FUNCTION "LGF_MatrixSubtraction" : Void   // FC10010, SCL
{ S7_Optimized_Access := 'TRUE' }
   VAR_INPUT
      matrix1 : Array[*, *] of Real;   // minuend
      matrix2 : Array[*, *] of Real;   // subtrahend
   END_VAR
   VAR_OUTPUT
      matrixResult : Array[*, *] of Real;   // result matrix
      error : Bool;
      statusID : UInt;
      status : Word;
   END_VAR
   VAR_TEMP
      tempMatrix1LowerBound1Dim : DInt;   // -
      tempMatrix1LowerBound2Dim : DInt;   // -
      tempMatrix1UpperBound1Dim : DInt;   // -
      tempMatrix1UpperBound2Dim : DInt;   // -
      tempMatrix2LowerBound1Dim : DInt;   // -
      tempMatrix2LowerBound2Dim : DInt;   // -
      tempMatrix2UpperBound1Dim : DInt;   // -
      tempMatrix2UpperBound2Dim : DInt;   // -
      tempResultMatrixLowerBound1Dim : DInt;   // -
      tempResultMatrixLowerBound2Dim : DInt;   // -
      tempResultMatrixUpperBound1Dim : DInt;   // -
      tempResultMatrixUpperBound2Dim : DInt;   // -
      tempCounterDim1 : Int;   // -
      tempCounterDim2 : Int;   // -
   END_VAR
   VAR CONSTANT
      NO_ERROR : Word := 16#0000;   // No errors.
      ERROR_LOWER_BOUND_NOT_EQUAL : Word := 16#8200;   // Lower bounds of matrices are not equal.
      ERROR_UPPER_BOUND_NOT_EQUAL : Word := 16#8201;   // Upper bounds of matrices are not equal.
      ERROR_IN_THIS_BLOCK : UInt := 1;   // statusID: Error in this block.
   END_VAR
BEGIN
   //=============================================================================
   // SIEMENS AG
   // (c)Copyright 2017
   //-----------------------------------------------------------------------------
   // Library:       LGF (Library General Functions)
   // Tested with:   CPU1212C DC/DC/DC FW:V4.2
   // Engineering:   TIA Portal V14 Update 1
   // Restrictions:  -
   // Requirements:  PLC (S7-1200 / S7-1500)
   // Functionality: This function subtracts matrices.
   //-----------------------------------------------------------------------------
   // Change log table:
   // Version  Date        In charge / Changes applied
   // 01.00.00 19.08.2015  Siemens Industry Online Support
   //                      First released version
   // 01.00.01 02.01.2017  Siemens Industry Online Support
   //                      Upgrade: TIA Portal V14 Update 1
   // 02.00.00 06.02.2017  Siemens Industry Online Support
   //                      Functionality using Array[*,*]
   // 02.00.01 17.08.2018  Siemens Industry Online Support
   //                      Upgrade: TIA V15 Update 2
   // 02.00.02 23.11.2018  Siemens Industry Online Support
   //                      Upgrade: TIA V15.1
   //=============================================================================

   //Set "No error" status
   #error := false;
   #statusID := #ERROR_IN_THIS_BLOCK;
   #status := #NO_ERROR;

   // Init resultMatrix
   #matrixResult[0, 0] := 0.0;

   //Determine the size of the matrices
   // Lower bound dimension 1
   #tempMatrix1LowerBound1Dim := LOWER_BOUND(ARR := #matrix1, DIM := 1);
   #tempMatrix2LowerBound1Dim := LOWER_BOUND(ARR := #matrix2, DIM := 1);
   #tempResultMatrixLowerBound1Dim := LOWER_BOUND(ARR := #matrixResult, DIM := 1);
   // Lower bound dimension 2
   #tempMatrix1LowerBound2Dim := LOWER_BOUND(ARR := #matrix1, DIM := 2);
   #tempMatrix2LowerBound2Dim := LOWER_BOUND(ARR := #matrix2, DIM := 2);
   #tempResultMatrixLowerBound2Dim := LOWER_BOUND(ARR := #matrixResult, DIM := 2);
   // Upper bound dimension 1
   #tempMatrix1UpperBound1Dim := UPPER_BOUND(ARR := #matrix1, DIM := 1);
   #tempMatrix2UpperBound1Dim := UPPER_BOUND(ARR := #matrix2, DIM := 1);
   #tempResultMatrixUpperBound1Dim := UPPER_BOUND(ARR := #matrixResult, DIM := 1);
   // Upper bound dimension 2
   #tempMatrix1UpperBound2Dim := UPPER_BOUND(ARR := #matrix1, DIM := 2);
   #tempMatrix2UpperBound2Dim := UPPER_BOUND(ARR := #matrix2, DIM := 2);
   #tempResultMatrixUpperBound2Dim := UPPER_BOUND(ARR := #matrixResult, DIM := 2);

   // Check the lower bound of all matrices
   IF (#tempMatrix1LowerBound1Dim <> #tempMatrix2LowerBound1Dim) OR (#tempMatrix1LowerBound1Dim <> #tempResultMatrixLowerBound1Dim) OR
     (#tempMatrix1LowerBound2Dim <> #tempMatrix2LowerBound2Dim) OR (#tempMatrix1LowerBound2Dim <> #tempResultMatrixLowerBound2Dim) THEN
     #error := TRUE;
     #status := #ERROR_LOWER_BOUND_NOT_EQUAL;
     RETURN;
   END_IF;
   // Check the upper bound of all matrices
   IF (#tempMatrix1UpperBound1Dim <> #tempMatrix2UpperBound1Dim) OR (#tempMatrix1UpperBound1Dim <> #tempResultMatrixUpperBound1Dim) OR
     (#tempMatrix1UpperBound2Dim <> #tempMatrix2UpperBound2Dim) OR (#tempMatrix1UpperBound2Dim <> #tempResultMatrixUpperBound2Dim) THEN
     #error := TRUE;
     #status := #ERROR_UPPER_BOUND_NOT_EQUAL;
     RETURN;
   END_IF;

   // Subtraction of two matrices
   FOR #tempCounterDim1 := #tempMatrix1LowerBound1Dim TO #tempMatrix1UpperBound1Dim DO
     FOR #tempCounterDim2 := #tempMatrix1LowerBound2Dim TO #tempMatrix1UpperBound2Dim DO
       #matrixResult[#tempCounterDim1, #tempCounterDim2] := #matrix1[#tempCounterDim1, #tempCounterDim2] - #matrix2[#tempCounterDim1, #tempCounterDim2];
     END_FOR;
   END_FOR;
END_FUNCTION

FUNCTION "LGF_MatrixTranspose" : Void   // FC10011, SCL
{ S7_Optimized_Access := 'TRUE' }
   VAR_INPUT
      matrix : Array[*, *] of Real;   // Matrix to be transposed.
   END_VAR
   VAR_OUTPUT
      matrixResult : Array[*, *] of Real;   // Transposed matrix.
      error : Bool;
      statusID : UInt;
      status : Word;
   END_VAR
   VAR_TEMP
      tempMatrixLowerBound1Dim : DInt;   // -
      tempMatrixLowerBound2Dim : DInt;   // -
      tempMatrixUpperBound1Dim : DInt;   // -
      tempMatrixUpperBound2Dim : DInt;   // -
      tempResultMatrixLowerBound1Dim : DInt;   // -
      tempResultMatrixLowerBound2Dim : DInt;   // -
      tempResultMatrixUpperBound1Dim : DInt;   // -
      tempResultMatrixUpperBound2Dim : DInt;   // -
      tempCounterDim1 : Int;   // -
      tempCounterDim2 : Int;   // -
   END_VAR
   VAR CONSTANT
      NO_ERROR : Word := 16#0000;   // No error.
      ERROR_LOWER_BOUND : Word := 16#8200;   // Lower bound of "matrixResult" is different to "matrix".
      ERROR_UPPER_BOUND : Word := 16#8201;   // Upper bound of "matrixResult" is different to "matrix".
      ERROR_IN_THIS_BLOCK : UInt := 1;   // statusID: Error in this block.
   END_VAR
BEGIN
   //=============================================================================
   // SIEMENS AG
   // (c)Copyright 2017
   //-----------------------------------------------------------------------------
   // Library:       LGF (Library General Functions)
   // Tested with:   CPU1212C DC/DC/DC FW:V4.2
   // Engineering:   TIA Portal V14 Update 1
   // Restrictions:  -
   // Requirements:  PLC (S7-1200 / S7-1500)
   // Functionality: This function transposes matrices.
   //-----------------------------------------------------------------------------
   // Change log table:
   // Version  Date        In charge / Changes applied
   // 01.00.00 19.08.2015  Siemens Industry Online Support
   //                      First released version
   // 01.00.01 02.01.2017  Siemens Industry Online Support
   //                      Upgrade: TIA Portal V14 Update 1
   // 02.00.00 06.02.2017  Siemens Industry Online Support
   //                      Functionality using Array[*,*]
   // 02.00.01 17.08.2018  Siemens Industry Online Support
   //                      Upgrade: TIA V15 Update 2
   // 02.00.02 23.11.2018  Siemens Industry Online Support
   //                      Upgrade: TIA V15.1
   //=============================================================================

   //Set "No error" status
   #error := false;
   #statusID := #ERROR_IN_THIS_BLOCK;
   #status := #NO_ERROR;

   // Init resultMatrix
   #matrixResult[0, 0] := 0.0;

   //Determine the size of the matrices
   // Lower bound dimension 1
   #tempMatrixLowerBound1Dim := LOWER_BOUND(ARR := #matrix, DIM := 1);
   #tempResultMatrixLowerBound1Dim := LOWER_BOUND(ARR := #matrixResult, DIM := 1);
   // Lower bound dimension 2
   #tempMatrixLowerBound2Dim := LOWER_BOUND(ARR := #matrix, DIM := 2);
   #tempResultMatrixLowerBound2Dim := LOWER_BOUND(ARR := #matrixResult, DIM := 2);
   // Upper bound dimension 1
   #tempMatrixUpperBound1Dim := UPPER_BOUND(ARR := #matrix, DIM := 1);
   #tempResultMatrixUpperBound1Dim := UPPER_BOUND(ARR := #matrixResult, DIM := 1);
   // Upper bound dimension 2
   #tempMatrixUpperBound2Dim := UPPER_BOUND(ARR := #matrix, DIM := 2);
   #tempResultMatrixUpperBound2Dim := UPPER_BOUND(ARR := #matrixResult, DIM := 2);

   // Check whether lower bounds of "matrixResult suit to the input "matrix"
   IF (#tempMatrixLowerBound1Dim <> #tempResultMatrixLowerBound2Dim) OR (#tempMatrixLowerBound2Dim <> #tempResultMatrixLowerBound1Dim) THEN
     #error := TRUE;
     #status := #ERROR_LOWER_BOUND;
     RETURN;
   END_IF;
   // Check whether upper bounds of "matrixResult suit to the input "matrix"
   IF (#tempMatrixUpperBound1Dim <> #tempResultMatrixUpperBound2Dim) OR (#tempMatrixUpperBound2Dim <> #tempResultMatrixUpperBound1Dim) THEN
     #error := TRUE;
     #status := #ERROR_UPPER_BOUND;
     RETURN;
   END_IF;

   //Transpose of the matrix
   FOR #tempCounterDim1 := #tempMatrixLowerBound1Dim TO #tempMatrixUpperBound1Dim DO
     FOR #tempCounterDim2 := #tempMatrixLowerBound2Dim TO #tempMatrixUpperBound2Dim DO
       #matrixResult[#tempCounterDim2, #tempCounterDim1] := #matrix[#tempCounterDim1, #tempCounterDim2];
     END_FOR;
   END_FOR;
END_FUNCTION

FUNCTION "LGF_RandomReal" : Real   // FC10014, SCL
{ S7_Optimized_Access := 'TRUE' }
   VAR_INPUT
      minValue : Real;   // minimal Value random can reach
      maxValue : Real;   // maximal Value random can reach
   END_VAR
   VAR_OUTPUT
      error : Bool;
      statusID : UInt;
      status : Word;
   END_VAR
   VAR_TEMP
      tempTime : DTL;
      tempTimeStatus : Int;
      tempRandomValue : UDInt;
      tempNormReal : Real;
   END_VAR
   VAR CONSTANT
      NO_ERROR : Word := 16#0000;
      NO_CURRENT_JOBS : Word := 16#7000;
      MAX_LESS_MIN : Word := 16#8200;
      ERROR_IN_THIS_BLOCK : UInt := 1;
      ERROR_RD_SYS_T : UInt := 2;
      MIN_UDINT : UDInt := 0;
      MAX_UDINT : UDInt := 4294967295;
   END_VAR
BEGIN
   //=============================================================================
   // Siemens AG
   // (c)Copyright 2017
   //-----------------------------------------------------------------------------
   // Library:       LGF (Library General Functions)
   // Tested with:   CPU1212C DC/DC/DC FW:V4.2
   // Engineering:   TIA Portal V14 Update 1
   // Restrictions:  -
   // Requirements:  PLC (S7-1200 / S7-1500)
   // Functionality: This function generates random numbers in defined limits
   //                (Datatype Real)
   //-----------------------------------------------------------------------------
   // Change log table:
   // Version  Date        In charge / Changes applied
   // 01.00.00 19.08.2015  Siemens Industry Online Support
   //                      First released version
   // 01.00.01 02.01.2017  Siemens Industry Online Support
   //                      Upgrade: TIA Portal V14 Update 1
   // 01.00.02 02.03.2017  Siemens Industry Online Support
   //                      Bugfix: FC number
   // 01.00.03 17.08.2018  Siemens Industry Online Support
   //                      Upgrade: TIA V15 Update 2
   // 01.00.04 23.11.2018  Siemens Industry Online Support
   //                      Upgrade: TIA V15.1
   //-----------------------------------------------------------------------------
   //Status Codes:
   // 16#7000:  No current jobs
   // 16#0000:  Job finished   // Note: There is no "Busy"-Status because the
   //           block is finished within a single cycle
   // 16#8200:  maxValue is samller then minValue 
   //=============================================================================

   //Set "No current job" status
   #error := false;
   #statusID := #ERROR_IN_THIS_BLOCK;
   #status := #NO_CURRENT_JOBS;

   //Check if the maximal Value is less than the minimal value
   IF (#minValue > #maxValue) THEN
     #error := true;
     #statusID := #ERROR_IN_THIS_BLOCK;
     #status := #MAX_LESS_MIN;
     #LGF_RandomReal := 0;
     RETURN;
   END_IF;

   //Read system time
   #tempTimeStatus := RD_SYS_T(#tempTime);

   IF (#tempTimeStatus <> 0) THEN
     #error := true;
     #statusID := #ERROR_RD_SYS_T;
     #status := INT_TO_WORD(#tempTimeStatus);
     #LGF_RandomReal := 0;
     RETURN;
   END_IF;

   //Callculate a random-start-value depending on the time
   #tempRandomValue.%B3 := #tempTime.NANOSECOND.%B0;
   #tempRandomValue.%B2 := #tempTime.NANOSECOND.%B1;
   #tempRandomValue.%B1 := #tempTime.NANOSECOND.%B2;
   #tempRandomValue.%B0 := #tempTime.NANOSECOND.%B3;

   //adapt the calculated random number to the given number span
   #tempNormReal := NORM_X(MIN := #MIN_UDINT, VALUE := #tempRandomValue, MAX := #MAX_UDINT);
   #LGF_RandomReal := SCALE_X(MIN := #minValue, VALUE := #tempNormReal, MAX := #maxValue);

   #status := #NO_ERROR;
END_FUNCTION

FUNCTION "LGF_SearchMinMax" : Void   // FC10015, SCL
{ S7_Optimized_Access := 'TRUE' }
   VAR_INPUT
      variableArray : Variant;
   END_VAR
   VAR_OUTPUT
      minValue : Variant;
      minArrayIndex : Int;
      maxValue : Variant;
      maxArrayIndex : Int;
      error : Bool;
      statusID : UInt;
      status : Word;
   END_VAR
   VAR_TEMP
      tempArraySize : UDInt;
      tempSizeCounter : Int;
      tempInternalError : Int;
      tempActValueInt : Int;
      tempMinInt : Int;
      tempArrayIndexMin : Int;
      tempMaxInt : Int;
      tempArrayIndexMax : Int;
      tempActValueUInt : UInt;
      tempMinUInt : UInt;
      tempMaxUInt : UInt;
      tempActValueDInt : DInt;
      tempMinDInt : DInt;
      tempMaxDInt : DInt;
      tempActValueUDInt : UDInt;
      tempMinUDInt : UDInt;
      tempMaxUDInt : UDInt;
      tempActValueUSInt : USInt;
      tempMinUSInt : USInt;
      tempMaxUSInt : USInt;
      tempActValueSInt : SInt;
      tempMinSInt : SInt;
      tempMaxSInt : SInt;
      tempActValueReal : Real;
      tempMinReal : Real;
      tempMaxReal : Real;
   END_VAR
   VAR CONSTANT
      NO_ERROR : Word := 16#0000;
      NO_CURRENT_JOBS : Word := 16#7000;
      NO_ARRAY : Word := 16#8200;
      WRONG_TYPE : Word := 16#8201;
      NOT_EQUAL_TYPES : Word := 16#8202;
      ERROR_IN_THIS_BLOCK : UInt := 1;
      ERROR_MOVE_BLK_VARIANT : UInt := 2;
   END_VAR
BEGIN
   //=============================================================================
   // SIEMENS AG
   // (c)Copyright 2017
   //-----------------------------------------------------------------------------
   // Library:       LGF (Library General Functions)
   // Tested with:   CPU1212C DC/DC/DC FW:V4.2
   // Engineering:   TIA Portal V14 Update 1
   // Restrictions:  -
   // Requirements:  PLC (S7-1200 / S7-1500)
   // Functionality: This function searches the min and max value in an array
   //-----------------------------------------------------------------------------
   // Change log table:
   // Version  Date        In charge / Changes applied
   // 01.00.00 19.08.2015  Siemens Industry Online Support
   //                      First released version
   // 01.00.01 02.01.2017  Siemens Industry Online Support
   //                      Upgrade: TIA Portal V14 Update 1
   // 01.00.02 17.08.2018  Siemens Industry Online Support
   //                      Upgrade: TIA V15 Update 2
   // 01.00.03 23.11.2018  Siemens Industry Online Support
   //                      Upgrade: TIA V15.1
   //=============================================================================

   // Set "No current job" status
   #error := false;
   #statusID := #ERROR_IN_THIS_BLOCK;
   #status := #NO_CURRENT_JOBS;
   #tempInternalError := 0;

   // Check if the variant-variable is an array if yes cout the elements of the array
   IF NOT (IS_ARRAY(#variableArray)) THEN
     #error := true;
     #statusID := #ERROR_IN_THIS_BLOCK;
     #status := #NO_ARRAY;
     RETURN;
   ELSE
     #tempArraySize := CountOfElements(#variableArray);
   END_IF;

   // Check if the elements of the array and the variables min and max have the same datatype.
   IF TypeOfElements(#variableArray) <> TypeOf(#minValue) OR TypeOf(#minValue) <> TypeOf(#maxValue) THEN
     #error := true;
     #statusID := #ERROR_IN_THIS_BLOCK;
     #status := #NOT_EQUAL_TYPES;
     RETURN;
   END_IF;

   //Request of the datatype
   CASE TypeOfElements(#variableArray) OF
     Int:
       //----------------------- Search min -------------------------------
       #tempMinInt := 32767;
       FOR #tempSizeCounter := 0 TO UDINT_TO_INT(#tempArraySize) DO

         //Read the next element of the array
         #tempInternalError := MOVE_BLK_VARIANT(SRC := #variableArray,
                                                COUNT := 1,
                                                SRC_INDEX := #tempSizeCounter,
                                                DEST_INDEX := 0,
                                                DEST => #tempActValueInt);

         //compare the new value with the actual best value
         IF #tempActValueInt < #tempMinInt THEN
           #tempMinInt := #tempActValueInt;
           #tempArrayIndexMin := #tempSizeCounter;
         END_IF;

       END_FOR;

       //copy the data to the outputs
       #minArrayIndex := #tempArrayIndexMin;
       #tempInternalError := MOVE_BLK_VARIANT(SRC := #tempMinInt,
                                              COUNT := 1,
                                              SRC_INDEX := 0,
                                              DEST_INDEX := 0,
                                              DEST => #minValue);

       //----------------------- Search max -------------------------------
       #tempMaxInt := -32768;
       FOR #tempSizeCounter := 0 TO UDINT_TO_INT(#tempArraySize) DO

         //Read the next element of the array
         #tempInternalError := MOVE_BLK_VARIANT(SRC := #variableArray,
                                                COUNT := 1,
                                                SRC_INDEX := #tempSizeCounter,
                                                DEST_INDEX := 0,
                                                DEST => #tempActValueInt);

         //compare the new value with the actual best value
         IF #tempActValueInt > #tempMaxInt THEN
           #tempMaxInt := #tempActValueInt;
           #tempArrayIndexMax := #tempSizeCounter;
         END_IF;

       END_FOR;

       //copy the data to the outputs
       #maxArrayIndex := #tempArrayIndexMax;
       #tempInternalError := MOVE_BLK_VARIANT(SRC := #tempMaxInt,
                                              COUNT := 1,
                                              SRC_INDEX := 0,
                                              DEST_INDEX := 0,
                                              DEST => #maxValue);

     UInt:
       //----------------------- Search min -------------------------------
       #tempMinUInt := 65535;
       FOR #tempSizeCounter := 0 TO UDINT_TO_INT(#tempArraySize) DO

         //Read the next element of the array
         #tempInternalError := MOVE_BLK_VARIANT(SRC := #variableArray,
                                                COUNT := 1,
                                                SRC_INDEX := #tempSizeCounter,
                                                DEST_INDEX := 0,
                                                DEST => #tempActValueUInt);

         //compare the new value with the actual best value
         IF #tempActValueUInt < #tempMinUInt THEN
           #tempMinUInt := #tempActValueUInt;
           #tempArrayIndexMin := #tempSizeCounter;
         END_IF;

       END_FOR;

       //copy the data to the outputs
       #minArrayIndex := #tempArrayIndexMin;
       #tempInternalError := MOVE_BLK_VARIANT(SRC := #tempMinUInt,
                                              COUNT := 1,
                                              SRC_INDEX := 0,
                                              DEST_INDEX := 0,
                                              DEST => #minValue);

       //----------------------- Search max -------------------------------
       #tempMaxUInt := 0;
       FOR #tempSizeCounter := 0 TO UDINT_TO_INT(#tempArraySize) DO

         //Read the next element of the array
         #tempInternalError := MOVE_BLK_VARIANT(SRC := #variableArray,
                                                COUNT := 1,
                                                SRC_INDEX := #tempSizeCounter,
                                                DEST_INDEX := 0,
                                                DEST => #tempActValueUInt);

         //compare the new value with the actual best value
         IF #tempActValueUInt > #tempMaxUInt THEN
           #tempMaxUInt := #tempActValueUInt;
           #tempArrayIndexMax := #tempSizeCounter;
         END_IF;

       END_FOR;

       //copy the data to the outputs
       #maxArrayIndex := #tempArrayIndexMax;
       #tempInternalError := MOVE_BLK_VARIANT(SRC := #tempMaxUInt,
                                              COUNT := 1,
                                              SRC_INDEX := 0,
                                              DEST_INDEX := 0,
                                              DEST => #maxValue);

     DInt:
       //----------------------- Search min -------------------------------
       #tempMinDInt := 2147483647;
       FOR #tempSizeCounter := 0 TO UDINT_TO_INT(#tempArraySize) DO

         #tempInternalError := MOVE_BLK_VARIANT(SRC := #variableArray,
                                                COUNT := 1,
                                                SRC_INDEX := #tempSizeCounter,
                                                DEST_INDEX := 0,
                                                DEST => #tempActValueDInt);
         IF #tempActValueDInt < #tempMinDInt THEN
           #tempMinDInt := #tempActValueDInt;
           #tempArrayIndexMin := #tempSizeCounter;
         END_IF;

       END_FOR;

       #minArrayIndex := #tempArrayIndexMin;
       #tempInternalError := MOVE_BLK_VARIANT(SRC := #tempMinDInt,
                                              COUNT := 1,
                                              SRC_INDEX := 0,
                                              DEST_INDEX := 0,
                                              DEST => #minValue);

       //----------------------- Search max -------------------------------
       #tempMaxDInt := -2147483648;
       FOR #tempSizeCounter := 0 TO UDINT_TO_INT(#tempArraySize) DO

         #tempInternalError := MOVE_BLK_VARIANT(SRC := #variableArray,
                                                COUNT := 1,
                                                SRC_INDEX := #tempSizeCounter,
                                                DEST_INDEX := 0,
                                                DEST => #tempActValueDInt);
         IF #tempActValueDInt > #tempMaxDInt THEN
           #tempMaxDInt := #tempActValueDInt;
           #tempArrayIndexMax := #tempSizeCounter;
         END_IF;

       END_FOR;

       #maxArrayIndex := #tempArrayIndexMax;
       #tempInternalError := MOVE_BLK_VARIANT(SRC := #tempMaxDInt,
                                              COUNT := 1,
                                              SRC_INDEX := 0,
                                              DEST_INDEX := 0,
                                              DEST => #maxValue);

     UDInt:
       //----------------------- Search min -------------------------------
       #tempMinUDInt := 4294967295;
       FOR #tempSizeCounter := 0 TO UDINT_TO_INT(#tempArraySize) DO

         #tempInternalError := MOVE_BLK_VARIANT(SRC := #variableArray,
                                                COUNT := 1,
                                                SRC_INDEX := #tempSizeCounter,
                                                DEST_INDEX := 0,
                                                DEST => #tempActValueUDInt);
         IF #tempActValueUDInt < #tempMinUDInt THEN
           #tempMinUDInt := #tempActValueUDInt;
           #tempArrayIndexMin := #tempSizeCounter;
         END_IF;

       END_FOR;

       #minArrayIndex := #tempArrayIndexMin;
       #tempInternalError := MOVE_BLK_VARIANT(SRC := #tempMinUDInt,
                                              COUNT := 1,
                                              SRC_INDEX := 0,
                                              DEST_INDEX := 0,
                                              DEST => #minValue);

       //----------------------- Search max -------------------------------
       #tempMaxUDInt := 0;
       FOR #tempSizeCounter := 0 TO UDINT_TO_INT(#tempArraySize) DO

         #tempInternalError := MOVE_BLK_VARIANT(SRC := #variableArray,
                                                COUNT := 1,
                                                SRC_INDEX := #tempSizeCounter,
                                                DEST_INDEX := 0,
                                                DEST => #tempActValueUDInt);
         IF #tempActValueUDInt > #tempMaxUDInt THEN
           #tempMaxUDInt := #tempActValueUDInt;
           #tempArrayIndexMax := #tempSizeCounter;
         END_IF;

       END_FOR;

       #maxArrayIndex := #tempArrayIndexMax;
       #tempInternalError := MOVE_BLK_VARIANT(SRC := #tempMaxUDInt,
                                              COUNT := 1,
                                              SRC_INDEX := 0,
                                              DEST_INDEX := 0,
                                              DEST => #maxValue);

     USInt:
       //----------------------- Search min -------------------------------
       #tempMinUSInt := 255;
       FOR #tempSizeCounter := 0 TO UDINT_TO_INT(#tempArraySize) DO

         #tempInternalError := MOVE_BLK_VARIANT(SRC := #variableArray,
                                                COUNT := 1,
                                                SRC_INDEX := #tempSizeCounter,
                                                DEST_INDEX := 0,
                                                DEST => #tempActValueUSInt);
         IF #tempActValueUSInt < #tempMinUSInt THEN
           #tempMinUSInt := #tempActValueUSInt;
           #tempArrayIndexMin := #tempSizeCounter;
         END_IF;

       END_FOR;

       #minArrayIndex := #tempArrayIndexMin;
       #tempInternalError := MOVE_BLK_VARIANT(SRC := #tempMinUSInt,
                                              COUNT := 1,
                                              SRC_INDEX := 0,
                                              DEST_INDEX := 0,
                                              DEST => #minValue);

       //----------------------- Search max -------------------------------
       #tempMaxUSInt := 0;
       FOR #tempSizeCounter := 0 TO UDINT_TO_INT(#tempArraySize) DO

         #tempInternalError := MOVE_BLK_VARIANT(SRC := #variableArray,
                                                COUNT := 1,
                                                SRC_INDEX := #tempSizeCounter,
                                                DEST_INDEX := 0,
                                                DEST => #tempActValueUSInt);
         IF #tempActValueUSInt > #tempMaxUSInt THEN
           #tempMaxUSInt := #tempActValueUSInt;
           #tempArrayIndexMax := #tempSizeCounter;
         END_IF;

       END_FOR;

       #maxArrayIndex := #tempArrayIndexMax;
       #tempInternalError := MOVE_BLK_VARIANT(SRC := #tempMaxUSInt,
                                              COUNT := 1,
                                              SRC_INDEX := 0,
                                              DEST_INDEX := 0,
                                              DEST => #maxValue);

     SInt:
       //----------------------- Search min -------------------------------
       #tempMinSInt := 127;
       FOR #tempSizeCounter := 0 TO UDINT_TO_INT(#tempArraySize) DO

         #tempInternalError := MOVE_BLK_VARIANT(SRC := #variableArray,
                                                COUNT := 1,
                                                SRC_INDEX := #tempSizeCounter,
                                                DEST_INDEX := 0,
                                                DEST => #tempActValueSInt);
         IF #tempActValueSInt < #tempMinSInt THEN
           #tempMinSInt := #tempActValueSInt;
           #tempArrayIndexMin := #tempSizeCounter;
         END_IF;

       END_FOR;

       #minArrayIndex := #tempArrayIndexMin;
       #tempInternalError := MOVE_BLK_VARIANT(SRC := #tempMinSInt,
                                              COUNT := 1,
                                              SRC_INDEX := 0,
                                              DEST_INDEX := 0,
                                              DEST => #minValue);

       //----------------------- Search max -------------------------------
       #tempMaxSInt := -128;
       FOR #tempSizeCounter := 0 TO UDINT_TO_INT(#tempArraySize) DO

         #tempInternalError := MOVE_BLK_VARIANT(SRC := #variableArray,
                                                COUNT := 1,
                                                SRC_INDEX := #tempSizeCounter,
                                                DEST_INDEX := 0,
                                                DEST => #tempActValueSInt);
         IF #tempActValueSInt > #tempMaxSInt THEN
           #tempMaxSInt := #tempActValueSInt;
           #tempArrayIndexMax := #tempSizeCounter;
         END_IF;

       END_FOR;

       #maxArrayIndex := #tempArrayIndexMax;
       #tempInternalError := MOVE_BLK_VARIANT(SRC := #tempMaxSInt,
                                              COUNT := 1,
                                              SRC_INDEX := 0,
                                              DEST_INDEX := 0,
                                              DEST => #maxValue);
     Real:
       //----------------------- Search min -------------------------------
       #tempInternalError := MOVE_BLK_VARIANT(SRC := #variableArray,
                                              COUNT := 1,
                                              SRC_INDEX := 0,
                                              DEST_INDEX := 0,
                                              DEST => #tempMinReal);

       FOR #tempSizeCounter := 0 TO UDINT_TO_INT(#tempArraySize) DO

         #tempInternalError := MOVE_BLK_VARIANT(SRC := #variableArray,
                                                COUNT := 1,
                                                SRC_INDEX := #tempSizeCounter,
                                                DEST_INDEX := 0,
                                                DEST => #tempActValueReal);
         IF #tempActValueReal < #tempMinReal THEN
           #tempMinReal := #tempActValueReal;
           #tempArrayIndexMin := #tempSizeCounter;
         END_IF;

       END_FOR;

       #minArrayIndex := #tempArrayIndexMin;
       #tempInternalError := MOVE_BLK_VARIANT(SRC := #tempMinReal,
                                              COUNT := 1,
                                              SRC_INDEX := 0,
                                              DEST_INDEX := 0,
                                              DEST => #minValue);

       //----------------------- Search max -------------------------------
       #tempInternalError := MOVE_BLK_VARIANT(SRC := #variableArray,
                                              COUNT := 1,
                                              SRC_INDEX := 0,
                                              DEST_INDEX := 0,
                                              DEST => #tempMaxReal);

       FOR #tempSizeCounter := 0 TO UDINT_TO_INT(#tempArraySize) DO

         #tempInternalError := MOVE_BLK_VARIANT(SRC := #variableArray,
                                                COUNT := 1,
                                                SRC_INDEX := #tempSizeCounter,
                                                DEST_INDEX := 0,
                                                DEST => #tempActValueReal);
         IF #tempActValueReal > #tempMaxReal THEN
           #tempMaxReal := #tempActValueReal;
           #tempArrayIndexMax := #tempSizeCounter;
         END_IF;

       END_FOR;

       #maxArrayIndex := #tempArrayIndexMax;
       #tempInternalError := MOVE_BLK_VARIANT(SRC := #tempMaxReal,
                                              COUNT := 1,
                                              SRC_INDEX := 0,
                                              DEST_INDEX := 0,
                                              DEST => #maxValue);
     ELSE
       #error := true;
       #statusID := #ERROR_IN_THIS_BLOCK;
       #status := #WRONG_TYPE;
       RETURN;
   END_CASE;

   IF #tempInternalError <> 0 THEN
     #error := true;
     #statusID := #ERROR_MOVE_BLK_VARIANT;
     #status := INT_TO_WORD(#tempInternalError);
     RETURN;
   END_IF;

   #status := #NO_ERROR;
END_FUNCTION

FUNCTION "LGF_XRoot" : Real   // FC10016, SCL
{ S7_Optimized_Access := 'TRUE' }
   VAR_INPUT
      variable : Real;   // To be extracted value. / Time value to convert
      root : Real;   // exponent of root / Execute Template
   END_VAR
   // Ret_Val : result of calculation / reset signal, rising edge
   VAR CONSTANT
      ONE : Real := 1.0;
   END_VAR
BEGIN
   //=============================================================================
   // SIEMENS AG
   // (c)Copyright 2017
   //-----------------------------------------------------------------------------
   // Library:       LGF (Library General Functions)
   // Tested with:   CPU1212C DC/DC/DC FW:V4.2
   // Engineering:   TIA Portal V14 Update 14
   // Restrictions:  -
   // Requirements:  PLC (S7-1200 / S7-1500)
   // Functionality: This function extracts a root.
   //-----------------------------------------------------------------------------
   // Change log table:
   // Version  Date        In charge / Changes applied
   // 01.00.00 19.08.2015  Siemens Industry Online Support
   //                      First released version
   // 01.00.01 02.01.2017  Siemens Industry Online Support
   //                      Upgrade: TIA Portal V14 Update 1
   // 01.00.02 17.08.2018  Siemens Industry Online Support
   //                      Upgrade: TIA V15 Update 2
   // 01.00.03 23.11.2018  Siemens Industry Online Support
   //                      Upgrade: TIA V15.1
   // 01.00.04 17.01.2019  Siemens Industry Online Support
   //                      Calculation changed
   //=============================================================================

   // Calculation of the x-th root
   #LGF_XRoot := #variable ** (#ONE / #root);
END_FUNCTION

FUNCTION "LGF_Distance" : LReal   // FC10020, SCL
{ S7_Optimized_Access := 'TRUE' }
VERSION : 0.1
   VAR_INPUT
      x1 : LReal;   // X coordinate point 1
      y1 : LReal;   // Y coordinate point 1
      x2 : LReal;   // X coordinate point 2
      y2 : LReal;   // Y coordinate point 2
   END_VAR
   VAR_TEMP
      tempXq : LReal;   // Square of difference X
      tempYq : LReal;   // Square of difference X
      tempDistance : LReal;   // Temporary calculated distance
   END_VAR
   // Ret_Val : Calculated distance
BEGIN
   //=============================================================================
   // Siemens AG
   // (c)Copyright 2017
   //-----------------------------------------------------------------------------
   // Library:       LGF (Library General Functions)
   // Tested with:   CPU1212C DC/DC/DC FW:V4.2
   // Engineering:   TIA Portal V15 Upd 2
   // Restrictions:  -
   // Requirements:  PLC (S7-1200 / S7-1500)
   // Functionality: This function calculates the distance between two points in
   //                a Cartesian coordinate system 
   //-----------------------------------------------------------------------------
   // Change log table:
   // Version  Date        In charge/Changes applied
   // 01.00.00 06.07.2018  Siemens Industry Online Support
   //                      First released version
   // 01.00.01 17.08.2018  Siemens Industry Online Support
   //                      Upgrade: TIA V15 Update 2
   // 01.00.02 23.11.2018  Siemens Industry Online Support
   //                      Upgrade: TIA V15.1
   // 01.01.00 25.01.2019  Siemens Industry Online Support
   //                      Data type changed to LREAL
   //-----------------------------------------------------------------------------
   //Status Codes: -
   //=============================================================================

   #tempDistance := 0;

   #tempXq := SQR(#x2 - #x1);
   #tempYq := SQR(#y2 - #y1);

   #tempDistance := SQRT(#tempXq + #tempYq);

   #LGF_Distance := #tempDistance;
END_FUNCTION

FUNCTION "LGF_RandomBasic" : Real   // FC10038, SCL
{ S7_Optimized_Access := 'TRUE' }
   VAR_TEMP
      tempTime : DTL;   // System time
      tempTimeStatus : Int;   // Status of the instruction RD_SYS_T
      tempRandomValue : UDInt;   // Random-start-value
   END_VAR
   // Ret_Val : Ret_Val
   VAR CONSTANT
      MIN_UDINT : UDInt := 0;   // UDInt lower value range
      MAX_UDINT : UDInt := 4294967295;   // UDInt upper value range
   END_VAR
BEGIN
   //=============================================================================
   // Siemens AG
   // (c)Copyright 2017
   //-----------------------------------------------------------------------------
   // Library:       LGF (Library General Functions)
   // Tested with:   CPU1212C DC/DC/DC FW:V4.2
   // Engineering:   TIA Portal V14 Upd 1
   // Restrictions:  -
   // Requirements:  PLC (S7-1200 / S7-1500)
   // Functionality: This function generates random numbers. 0.0 <= REAL <= 1.0
   //                (Datatype Real)
   //-----------------------------------------------------------------------------
   // Change log table:
   // Version  Date        In charge/Changes applied
   // 01.00.00 27.01.2017  Siemens Industry Online Support
   //                      First released version
   // 01.00.01 17.08.2018  Siemens Industry Online Support
   //                      Upgrade: TIA V15 Update 2
   // 01.00.02 23.11.2018  Siemens Industry Online Support
   //                      Upgrade: TIA V15.1
   //-----------------------------------------------------------------------------
   //Status Codes: -
   //=============================================================================

   //Read system time
   #tempTimeStatus := RD_SYS_T(#tempTime);

   //Callculate a random-start-value depending on the time
   #tempRandomValue.%B3 := #tempTime.NANOSECOND.%B0;
   #tempRandomValue.%B2 := #tempTime.NANOSECOND.%B1;
   #tempRandomValue.%B1 := #tempTime.NANOSECOND.%B2;
   #tempRandomValue.%B0 := #tempTime.NANOSECOND.%B3;

   //Norm the calculated random number: 0.0 <= #LGF_RandomBasic <= 1.0
   #LGF_RandomBasic := NORM_X(MIN := #MIN_UDINT, VALUE := #tempRandomValue, MAX := #MAX_UDINT);
END_FUNCTION

FUNCTION "LGF_HighLowLimit" : Void   // FC10040, SCL
{ S7_Optimized_Access := 'TRUE' }
VERSION : 0.1
   VAR_INPUT
      value : Real;   // Value to check if in deadband of setpoint
      setpoint : Real;   // Setpoint
      deadband : Real;   // Deadband
   END_VAR
   VAR_OUTPUT
      valueInRange : Bool;   // value is in range of the setpoint (deadband)
      valueOverHighLimit : Bool;   // value is over high limit
      valueUnderLowLimit : Bool;   // value is under low limit
      error : Bool;   // error
      status : Word;   // status
   END_VAR
   VAR_TEMP
      tempHighLimit : Real;   // Calculated high limit
      tempLowLimit : Real;   // Calculated low limit
      tempValueOverHighLimit : Bool;
      tempValueUnderLowLimit : Bool;
   END_VAR
   VAR CONSTANT
      NO_ERROR : Word := 16#0000;   // Status no error
      NO_CURRENT_JOBS : Word := 16#7000;   // -
      WRONG_VALUE_RANGE_HIGH_VALUE : Word := 16#8101;   // Status wrong value range high value
      WRONG_VALUE_RANGE_LOW_VALUE : Word := 16#8102;   // Status wrong value range low value
      MAX_LESS_MIN : Word := 16#8200;   // Status HighValue is smaller then LowValue -> error
      MAX_REAL_OVERFLOW : Real := 16#7F80_0000;   // Max Real value overflow
      MIN_REAL_OVERFLOW : Real := 16#FF80_0000;   // Min Real value overflow
   END_VAR
BEGIN
   //=============================================================================
   // Siemens AG
   // (c)Copyright 2017
   //-----------------------------------------------------------------------------
   // Library:       LGF (Library General Functions)
   // Tested with:   CPU1212C DC/DC/DC FW:V4.2
   // Engineering:   TIA Portal V14 Upd 1
   // Restrictions:  -
   // Requirements:  PLC (S7-1200 / S7-1500)
   // Functionality: This program calculates the low and high limit values
   //-----------------------------------------------------------------------------
   // Change log table:
   // Version  Date        In charge / Changes applied
   // 01.00.00 30.01.2017  Siemens Industry Online Support
   //                      First released version
   // 01.00.01 17.08.2018  Siemens Industry Online Support
   //                      Upgrade: TIA V15 Update 2
   // 01.00.02 23.11.2018  Siemens Industry Online Support
   //                      Upgrade: TIA V15.1
   //-----------------------------------------------------------------------------
   //Status Codes:
   // 16#0000:  Job finished   // Note: There is no "Busy"-Status because the
   //           block is finished within a single cycle
   // 16#8101:  Outside value range high value
   // 16#8102:  Outside value range low value
   // 16#8200:  highValue is samller then lowValue 
   //=============================================================================
   #error := FALSE;
   #status := #NO_CURRENT_JOBS;

   // Determination of high limit
   #tempHighLimit := #setpoint + (0.5 * ABS(#deadband));
   // Determination of low limit
   #tempLowLimit := #setpoint - (0.5 * ABS(#deadband));

   // High limit is smaller then LowValue -> error
   IF #tempHighLimit < #tempLowLimit THEN
     #error := TRUE;
     #status := #MAX_LESS_MIN;
     RETURN;
   END_IF;

   // Outside value data type range -> error
   IF (#tempHighLimit = #MAX_REAL_OVERFLOW) THEN
     #error := TRUE;
     #status := #WRONG_VALUE_RANGE_HIGH_VALUE;
     RETURN;
   ELSIF (#tempHighLimit = #MIN_REAL_OVERFLOW) THEN
     #error := TRUE;
     #status := #WRONG_VALUE_RANGE_HIGH_VALUE;
     RETURN;
   END_IF;

   IF (#tempLowLimit = #MAX_REAL_OVERFLOW) THEN
     #error := TRUE;
     #status := #WRONG_VALUE_RANGE_HIGH_VALUE;
     RETURN;
   ELSIF (#tempLowLimit = #MIN_REAL_OVERFLOW) THEN
     #error := TRUE;
     #status := #WRONG_VALUE_RANGE_LOW_VALUE;
     RETURN;
   END_IF;

   // Check if the value is higher then the high limit
   #tempValueOverHighLimit := #value > #tempHighLimit;

   // Check if the value is lower then the low limit
   #tempValueUnderLowLimit := #value < #tempLowLimit;

   // Check if the value is in range and write outputs
   #valueInRange := NOT (#tempValueOverHighLimit OR #tempValueUnderLowLimit);
   #valueOverHighLimit := #tempValueOverHighLimit;
   #valueUnderLowLimit := #tempValueUnderLowLimit;

   // No errors
   #status := #NO_ERROR;
END_FUNCTION

// folder: Phisical_functions/LGF/5 Data handling

FUNCTION_BLOCK "LGF_FIFO"   // FB10017, SCL
{ S7_Optimized_Access := 'TRUE' }
   VAR_INPUT
      execute : Bool;   // The instruction is executed when a positive signal edge is detected at the "request" parameter.
      mode : Bool;   // 0 = The first entry in the ring buffer is returned. 1 = An entry is written at the last position in the ring buffer.
      initialValue : Variant;   // Value with which the ARRAY of the ring buffer is initialized.
      resetBuffer : Bool;   // Clearing and initializing the buffer
   END_VAR
   VAR_OUTPUT
      error : Bool;   // Error
      statusID : UInt;   // Status ID
      status : Word;   // Status information
   END_VAR
   VAR_IN_OUT
      item : Variant;   // The entry that is either returned from the ring buffer or written to the ring buffer
      buffer : Variant;   // An ARRAY that is used as a ring buffer.
   END_VAR
   VAR
      statEdgeupm : Bool;   // Edge memory bit in which the RLO of the previous query is saved.
      statFirstItemIndex : Int := -1;   // Index of the oldest entry in the ring buffer
      statNextEmptyItemIndex : Int := 0;   // Index of the next free entry in the ring buffer
   END_VAR
   VAR_TEMP
      tempInternalError : Int;   // Error information
      tempNewFirstItemIndex : Int;   // Variable index
      tempNewNextEmptyItemIndex : Int;   // Variable index
      tempPufferSize : UDInt;   // Number of ARRAY elements in the ring buffer
      tempSizeCounter : Int;   // Size counter
   END_VAR
   VAR CONSTANT
      NO_ERROR : Word := 16#0000;   // No errors
      NO_CURRENT_JOBS : Word := 16#7000;   // Initial value
      BUFFER_EMPTY : Word := 16#8001;   // The buffer is empty
      BUFFER_FULL : Word := 16#8002;   // The buffer is full
      NO_ARRAY : Word := 16#8200;   // No array is present at the input "buffer"
      WRONG_TYPE_1 : Word := 16#8201;   // The data type of the InOut parameter "item" does not correspond to the data type of the array elements of the input "buffer"
      WRONG_TYPE_2 : Word := 16#8202;   // The data type of the input "initialValue" does not correspond to the data type of the InOut parameter "item"
      INDEX_IN_ARRAY_LIMITS_1 : Word := 16#8601;   // The tag "nextEmptyItemIndex" is not within the array limits
      INDEX_IN_ARRAY_LIMITS_2 : Word := 16#8602;   // The tag "firstItemIndex" is not within the array limits
      ERROR_IN_THIS_BLOCK : UInt := 1;   // Error in this block
      ERROR_MOVE_BLK_VARIANT : UInt := 2;   // Error/status of subordinate block "MOVE_BLK_VARIANT"
      NEXT_TASK_TO_EXECUTE : Bool := false;   // Next task to execute
      BUFFER_IS_EMPTY : Int := -1;   // Buffer is empty
      BUFFER_CONTAINS_ARRAY : Int := 0;   // Buffer contains array
      NO_INTERNAL_ERROR : Int := 0;   // No internal error
      BUFFER_INITIALIZED : Int := -1;   // Buffer initialized
      RESET : Bool := true;   // Reset
   END_VAR
BEGIN
   //=============================================================================
   // SIEMENS AG
   // (c)Copyright 2017
   //-----------------------------------------------------------------------------
   // Library:       LGF (Library General Functions)
   // Tested with:   CPU1212C DC/DC/DC FW:V4.2
   // Engineering:   TIA Portal V14
   // Restrictions:  -
   // Requirements:  PLC (S7-1200 / S7-1500)
   // Functionality: FIFO(First In First Out)-functionblock
   //-----------------------------------------------------------------------------
   // Change log table:
   // Version  Date        Expert in charge / Changes applied
   // 01.00.00 19.08.2015  Siemens Industry Online Support
   //                      First released version
   // 01.00.01 16.11.2015  Siemens Industry Online Support
   //                      Bug fix resetBuffer
   // 01.00.02 02.01.2017  Siemens Industry Online Support
   //                      Upgrade: TIA Portal V14 Update 1
   // 01.00.03 17.08.2018  Siemens Industry Online Support
   //                      Upgrade: TIA V15 Update 2
   // 01.00.04 23.11.2018  Siemens Industry Online Support
   //                      Upgrade: TIA V15.1
   // 02.00.00 29.01.2019  Siemens Industry Online Support
   //                      Output "done" removed (not necessary, because only one cycle)
   //=============================================================================

   //This program code section is only executed once after a negative signal edge.
   IF #execute = false AND #statEdgeupm = true THEN
     // If no error occurred during program execution, the error code "0000" is output.  
     #error := false;
     #statusID := #ERROR_IN_THIS_BLOCK;
     #status := #NO_CURRENT_JOBS;
   END_IF;

   //This program code section is only executed once after a positive signal edge.
   //IF there is no change in the signal state OF the result OF logic operation,
   //the program processing OF the "FIFOQueue" FB is terminated.

   IF #execute <> true OR #statEdgeupm <> false THEN
     #statEdgeupm := #execute;
     RETURN;
   END_IF;
   #statEdgeupm := #execute;

   // ------Validation of whether all parameter inputs are valid.----

   //This program code section checks whether the ring #buffer is an ARRAY.
   //IF so, the number OF the ARRAY elements is read out.
   //IF it is NOT an ARRAY, the program execution is terminated at this point
   //AND the status code "8200" is output.

   IF NOT (IS_ARRAY(#buffer)) THEN
     #error := true;
     #statusID := #ERROR_IN_THIS_BLOCK;
     #status := #NO_ARRAY;
     RETURN;
   ELSE
     #tempPufferSize := CountOfElements(#buffer);
   END_IF;

   //This program code section checks whether the data type OF the ARRAY elements matches
   //the data type OF the entry (tag #item). IF the data types DO NOT match,
   //the program execution is terminated at this point AND the error code "8201" is output.

   IF NOT (TypeOf(#item) = TypeOfElements(#buffer)) THEN
     #error := true;
     #statusID := #ERROR_IN_THIS_BLOCK;
     #status := #WRONG_TYPE_1;
     RETURN;
   END_IF;

   //This program code section checks whether the initial value OF the ring #buffer
   //matches the entry (tag #item). IF the data types DO NOT match,
   //the program execution is terminated at this point
   //AND the error code "8202" is output. *)

   IF NOT (TypeOf(#item) = TypeOf(#initialValue)) THEN
     #error := true;
     #statusID := #ERROR_IN_THIS_BLOCK;
     #status := #WRONG_TYPE_2;
     RETURN;
   END_IF;

   //This program code section checks whether the variable indices are within the ARRAY limits.
   //IF they are NOT, the program execution is terminated at this point
   //AND either error code "8601" OR "8602" is output depending on the index. *)

   IF (#statNextEmptyItemIndex >= #tempPufferSize) THEN
     #error := true;
     #statusID := #ERROR_IN_THIS_BLOCK;
     #status := #INDEX_IN_ARRAY_LIMITS_1;
     RETURN;
   END_IF;

   IF (#statFirstItemIndex >= #tempPufferSize) THEN
     #error := true;
     #statusID := #ERROR_IN_THIS_BLOCK;
     #status := #INDEX_IN_ARRAY_LIMITS_2;
     RETURN;
   END_IF;


   //If reset is "TRUE" the buffer and their  counters are resetted
   IF #resetBuffer = #RESET THEN
     #statFirstItemIndex := -1;
     #statNextEmptyItemIndex := 0;

     FOR #tempSizeCounter := 0 TO UDINT_TO_INT(#tempPufferSize - 1) DO

